// TIA Portal project "MCP_RB001002" (V15.1)

(* hardware
DEVICE "S7-1200 station_1"  S7-1200 Station
   slot 0: "Rack_0"  S7-1200 Rack  Rack  V1.0
   slot 1: "MCP"  CPU 1215C DC/DC/DC  6ES7 215-1AG40-0XB0  V4.2
DEVICE "GSD device_1"  GSD.Device.PN
   slot 0: "机架"  Rack  V1.0
   slot 0: "PNMB-address"  PNM02 V1.5  PNMB  V1.50
      slot 0: "PNM02 V1.5"  PNM02 V1.5
      slot 1: "PN-IO"  PN-IO
         slot 1: "Port 1"  Port 1
         slot 2: "Port 2"  Port 2
   slot 1: "M: 03 Read 050 Words (4xxxx)_1"  M: 03 Read 050 Words (4xxxx)
      slot 0: "M: 03 Read 050 Words (4xxxx)"  M: 03 Read 050 Words (4xxxx)
   slot 2: "M: 03 Read 050 Words (4xxxx)_2"  M: 03 Read 050 Words (4xxxx)
      slot 0: "M: 03 Read 050 Words (4xxxx)"  M: 03 Read 050 Words (4xxxx)
   slot 3: "M: 03 Read 050 Words (4xxxx)_3"  M: 03 Read 050 Words (4xxxx)
      slot 0: "M: 03 Read 050 Words (4xxxx)"  M: 03 Read 050 Words (4xxxx)
   slot 4: "M: 03 Read 050 Words (4xxxx)_4"  M: 03 Read 050 Words (4xxxx)
      slot 0: "M: 03 Read 050 Words (4xxxx)"  M: 03 Read 050 Words (4xxxx)
   slot 5: "M: 03 Read 050 Words (4xxxx)_5"  M: 03 Read 050 Words (4xxxx)
      slot 0: "M: 03 Read 050 Words (4xxxx)"  M: 03 Read 050 Words (4xxxx)
   slot 6: "M: 03 Read 002 Words (4xxxx)_1"  M: 03 Read 002 Words (4xxxx)
      slot 0: "M: 03 Read 002 Words (4xxxx)"  M: 03 Read 002 Words (4xxxx)
   slot 7: "M: 03 Read 002 Words (4xxxx)_2"  M: 03 Read 002 Words (4xxxx)
      slot 0: "M: 03 Read 002 Words (4xxxx)"  M: 03 Read 002 Words (4xxxx)
DEVICE "PC-System_1"  SIMATIC PC station
   slot 0: "SIMATIC PC station"  Rail  SIMATIC PC-Station  V1.0
      slot 125: "Stationmanager"  Station_Manager  V6.0.4
   slot 1: "IE general_1"  IE General  IE_CP  V8.2.0
   slot 2: "HMI_RT_1"  WinCC RT Advanced  6AV2 104-0xxxx-xxxx  15.1.0.0
      slot 33792: "主机接口"  Host interface
*)

// ===== PLC "MCP"  CPU 1215C DC/DC/DC =====

VAR_GLOBAL   // PLC tag table "默认变量表"
   "ID_100" AT %ID100 : Real;
   "ID_104" AT %ID104 : Real;
   "ID_108" AT %ID108 : Real;
   "ID_112" AT %ID112 : Real;
   "ID_116" AT %ID116 : Real;
   "ID_120" AT %ID120 : Real;
   "ID_124" AT %ID124 : Real;
   "ID_128" AT %ID128 : Real;
   "ID_132" AT %ID132 : Real;
   "ID_136" AT %ID136 : DInt;
   "ID_140" AT %ID140 : DInt;
   "ID_144" AT %ID144 : Real;
   "Tag_8" AT %ID148 : Real;
   "Tag_8(1)" AT %ID152 : Real;
   "Tag_9" AT %ID156 : Real;
   "ID_160" AT %IW160 : Word;
   "Tag_10" AT %ID164 : Real;
   "Tag_10(1)" AT %ID168 : Real;
   "Tag_11" AT %ID172 : Real;
   "Tag_11(1)" AT %ID176 : Real;
   "Tag_12" AT %ID180 : Real;
   "Tag_12(1)" AT %ID184 : Real;
   "Tag_13" AT %ID188 : Real;
   "Tag_13(1)" AT %ID192 : Real;
   "Tag_14" AT %ID196 : Real;
   "Tag_14(1)" AT %ID200 : Real;
   "Tag_15" AT %ID204 : Real;
   "Tag_16" AT %ID208 : Real;
   "Tag_17" AT %ID212 : Real;
   "Tag_18" AT %ID216 : Real;
   "Tag_19" AT %ID220 : Real;
   "Tag_20" AT %IW224 : Int;
   "Tag_21" AT %ID228 : Real;
   "Tag_22" AT %ID232 : Real;
   "Tag_23" AT %ID236 : Real;
   "Tag_24" AT %ID240 : Real;
   "Tag_25" AT %ID244 : Real;
   "Tag_26" AT %ID248 : Real;
   "Tag_27" AT %ID252 : Real;
   "Tag_28" AT %ID256 : Real;
   "Tag_29" AT %ID260 : Real;
   "Tag_30" AT %ID264 : Real;
   "Tag_31" AT %ID268 : Real;
   "Tag_32" AT %ID272 : Real;
   "Tag_33" AT %ID276 : Real;
   "ID_148" AT %ID148 : DWord;
   "ID_152" AT %ID152 : DWord;
   "ID_156" AT %ID156 : DWord;
   "ID_162" AT %IW162 : Word;
   "ID_164" AT %IW164 : Word;
   "ID_166" AT %IW166 : Word;
   "ID_168" AT %IW168 : Word;
   "ID_170" AT %IW170 : Word;
   "ID_172" AT %IW172 : Word;
   "ID_174" AT %IW174 : Word;
   "ID_176" AT %IW176 : Word;
   "ID_178" AT %IW178 : Word;
   "ID_180" AT %IW180 : Word;
   "ID_182" AT %IW182 : Word;
   "ID_184" AT %IW184 : Word;
   "ID_186" AT %IW186 : Word;
   "ID_188" AT %IW188 : Word;
   "ID_190" AT %IW190 : Word;
   "ID_192" AT %IW192 : Word;
   "ID_194" AT %IW194 : Word;
   "ID_196" AT %IW196 : Word;
   "ID_198" AT %IW198 : Word;
   "ID_158" AT %IW158 : Word;
   "Tag_1" AT %IW64 : Word;
   "Tag_2" AT %M100.0 : Bool;
   "Tag_3" AT %M100.1 : Bool;
   "Tag_4" AT %IW66 : Word;
   "Tag_5" AT %ID600 : DInt;
   "Tag_6" AT %ID700 : DInt;
   "Tag_7" AT %MD104 : DInt;
   "Tag_34" AT %MD108 : DInt;
   "System_Byte" AT %MB1 : Byte;
   "FirstScan" AT %M1.0 : Bool;
   "DiagStatusUpdate" AT %M1.1 : Bool;
   "AlwaysTRUE" AT %M1.2 : Bool;
   "AlwaysFALSE" AT %M1.3 : Bool;
   "Clock_Byte" AT %MB0 : Byte;
   "Clock_10Hz" AT %M0.0 : Bool;
   "Clock_5Hz" AT %M0.1 : Bool;
   "Clock_2.5Hz" AT %M0.2 : Bool;
   "Clock_2Hz" AT %M0.3 : Bool;
   "Clock_1.25Hz" AT %M0.4 : Bool;
   "Clock_1Hz" AT %M0.5 : Bool;
   "Clock_0.625Hz" AT %M0.6 : Bool;
   "Clock_0.5Hz" AT %M0.7 : Bool;
   "Tag_35" AT %M100.2 : Bool;
END_VAR

VAR_GLOBAL   // PLC tag table "精炼机采集"
   "N11" AT %I100.0 : "精炼机";
   "N12" AT %I200.0 : "精炼机";
   "N13" AT %I300.0 : "精炼机";
   "N14" AT %I400.0 : "精炼机";
   "N15" AT %I500.0 : "精炼机";
END_VAR

TYPE "精炼机"
   STRUCT
      左前辊温度 : Real;
      右前辊温度 : Real;
      左后辊温度 : Real;
      右后辊温度 : Real;
      左间隙 : Real;
      右间隙 : Real;
      滚筒电机电流 : Real;
      滚筒电机频率 : Real;
      滚筒电机功率 : Real;
      滚筒电机电度 : DInt;
      滚筒电机计时 : DInt;
      环境温度 : Real;
      环境湿度 : Real;
      胶温 : Real;
      开关量汇总 : DInt;
      当前任务编号 : Array[0..9] of WChar;
      当前人员编号 : Array[0..9] of WChar;
   END_STRUCT;
END_TYPE

TYPE "精炼机上传"
   STRUCT
      左前辊温度 : Real;
      右前辊温度 : Real;
      左后辊温度 : Real;
      右后辊温度 : Real;
      左间隙 : Real;
      右间隙 : Real;
      滚筒电机电流 : Real;
      滚筒电机频率 : Real;
      滚筒电机功率 : Real;
      滚筒电机电度 : DInt;
      滚筒电机计时 : DInt;
      环境温度 : Real;
      环境湿度 : Real;
      胶温 : Real;
      开关量汇总 : DInt;
      当前任务编号 : Array[0..9] of WChar;
      当前人员编号 : Array[0..9] of WChar;
   END_STRUCT;
END_TYPE

TYPE "uMySQL_CDD"
   STRUCT
      Connect_OK : Bool;
      Connect_ID : Conn_Ouc;
      Connect_Sequence : DInt;
      Server_Protocol_Version : Int;
      Server_Server_Version : String;
      Server_Character_Set : Byte;
      CLIENT_PLUGIN_AUTH : String;
      Recv_Done : Bool;
      Recv_Len : Int;
      Recv_Buffer : Array[0..2048] of Byte;
      Send_Done : Bool;
      Send_Len : Int;
      Send_Buffer : Array[0..2048] of Byte;
   END_STRUCT;
END_TYPE

TYPE "精炼机数据库"
   STRUCT
      左前辊温度 : Real;
      右前辊温度 : Real;
      左后辊温度 : Real;
      右后辊温度 : Real;
      左间隙 : Real;
      右间隙 : Real;
      滚筒电机电流 : Real;
      滚筒电机频率 : Real;
      滚筒电机功率 : Real;
      滚筒电机电度 : DInt;
      滚筒电机计时 : DInt;
      环境温度 : Real;
      环境湿度 : Real;
      胶温 : Real;
      开关量汇总 : DInt;
      当前任务编号 : WString;
      当前人员编号 : WString;
   END_STRUCT;
END_TYPE

DATA_BLOCK "精炼机数据转存"   // DB100
{ S7_Optimized_Access := 'FALSE' }
VERSION : 0.1
   VAR
      Temp : Array[0..99] of Byte;
      N11精炼机 : "精炼机上传";
      N12精炼机 : "精炼机上传";
      N13精炼机 : "精炼机上传";
      N14精炼机 : "精炼机上传";
      N15精炼机 : "精炼机上传";
      N21卷片机累计重量 : DInt;
      N22卷片机累计重量 : DInt;
   END_VAR
BEGIN
END_DATA_BLOCK

DATA_BLOCK "通用数据采集"   // DB200
{ S7_Optimized_Access := 'TRUE' }
VERSION : 0.1
   VAR
      环境温度 : Real;
      环境湿度 : Real;
   END_VAR
BEGIN
END_DATA_BLOCK

DATA_BLOCK "温控相机解码_N15"   // DB405
{ S7_Optimized_Access := 'TRUE' }
VERSION : 0.1
// stored: InstanceOfName 温控相机解码
"温控相机解码"
BEGIN
END_DATA_BLOCK

// folder: System blocks/Program resources

DATA_BLOCK "IEC_Timer_0_DB"   // DB1
{ S7_Optimized_Access := 'TRUE' }
AUTHOR : Simatic
FAMILY : IEC
NAME : IEC_TMR
VERSION : 1.0
// stored: InstanceOfName IEC_TIMER
"IEC_TIMER"
BEGIN
END_DATA_BLOCK

// folder: 存数据库

DATA_BLOCK "Wchartest"   // DB2
{ S7_Optimized_Access := 'TRUE' }
VERSION : 0.1
   VAR
      TemWchar : WChar;
      TemWstring : WString;
      WstringLen : UInt;
      ArrayWCHAR : Array[0..1023] of WChar;
      ArrayChar : Array[0..1023] of Char;
      arraayWord : Array[0..1023] of Word;
   END_VAR
BEGIN
END_DATA_BLOCK

DATA_BLOCK "数据库字符串"   // DB900
{ S7_Optimized_Access := 'TRUE' }
VERSION : 0.1
   VAR
      wstring : WString[2048];
   END_VAR
   VAR RETAIN
      Connect_CMD : Bool;
   END_VAR
   VAR
      Connect_CND : Bool;
      Connect_Error : Bool;
      Use_CMD : Bool;
      Use_Done : Bool;
      Use_Error : Bool;
      Query_CMD : Bool;
      Query_Done : Bool;
      Query_Error : Bool;
      CommandLine : WString[2048];
   END_VAR
   VAR RETAIN
      SerialNum : Int := 1;
   END_VAR
   VAR
      Addr : Int := 11;
      UploadData : "精炼机数据库";
      Upload : Array[11..15] of "精炼机数据库";
   END_VAR
BEGIN
END_DATA_BLOCK

DATA_BLOCK "uMySQL_Connect_DB"   // DB901
{ S7_Optimized_Access := 'TRUE' }
VERSION : 0.1
// stored: InstanceOfName uMySQL_Connect
"uMySQL_Connect"
BEGIN
   IP.RemoteAddress.ADDR[3] := 16#A0;
   IP.RemoteAddress.ADDR[4] := 16#A3;
   Net_ID := 16#0070;
   UserName := 'plc';
   DB_Name := 'rb001011';
   IP.InterfaceId := 64;
   IP.ID := 16#0070;
   IP.ConnectionType := 16#0B;
   IP.ActiveEstablished := TRUE;
   TempBool[1] := TRUE;
   SND_Buffer[0] := 16#01;
   SND_Buffer[4] := 16#01;
   NetConnect.STATUS := 16#7000;
   NetRcv.ADHOC := TRUE;
   NetRcv.STATUS := 16#7000;
   "Step" := 6;
   ServerCapability_flag := 16#0000_0000;
   Client_CapabilityFlag := 16#0000_8609;
   Client_MaxLen := 16#0000_0000;
   NetDISCON.ID := 16#0070;
   NetDISCON.STATUS := 16#7000;
   NetSend.ID := 16#0070;
   NetSend.STATUS := 16#7000;
   NetDiag.REQ := TRUE;
   NetDiag.ID := 16#0070;
   NetDiag.BUSY := TRUE;
   NetDiag.STATUS := 16#7001;
   Timer_ON.ST := T#10D_22H_43M_20S_90MS;
   Timer_ON.PT := T#500MS;
   Timer_ON.RU := TRUE;
   Timer_ON.IN := TRUE;
   Timer_OFF.ST := T#10D_22H_43M_19S_563MS;
   Timer_OFF.PT := T#500MS;
   NetSendEnd.REQ := TRUE;
   NetSendEnd.ID := 16#0070;
   NetSendEnd.LEN := 5;
   NetSendEnd.STATUS := 16#7000;
   NetSendEnd_EN := TRUE;
   SendWChar[0] := WCHAR#' ';
   SendWChar[1] := WCHAR#' ';
   SendWChar[2] := WCHAR#' ';
   SendWChar[3] := WCHAR#' ';
   SendWChar[4] := WCHAR#' ';
   SendWChar[5] := WCHAR#' ';
   SendWChar[6] := WCHAR#' ';
   SendWChar[7] := WCHAR#' ';
   SendWChar[8] := WCHAR#' ';
   SendWChar[9] := WCHAR#' ';
   SendWChar[10] := WCHAR#' ';
   SendWChar[11] := WCHAR#' ';
   SendWChar[12] := WCHAR#' ';
   SendWChar[13] := WCHAR#' ';
   SendWChar[14] := WCHAR#' ';
   SendWChar[15] := WCHAR#' ';
   SendWChar[16] := WCHAR#' ';
   SendWChar[17] := WCHAR#' ';
   SendWChar[18] := WCHAR#' ';
   SendWChar[19] := WCHAR#' ';
   SendWChar[20] := WCHAR#' ';
   SendWChar[21] := WCHAR#' ';
   SendWChar[22] := WCHAR#' ';
   SendWChar[23] := WCHAR#' ';
   SendWChar[24] := WCHAR#' ';
   SendWChar[25] := WCHAR#' ';
   SendWChar[26] := WCHAR#' ';
   SendWChar[27] := WCHAR#' ';
   SendWChar[28] := WCHAR#' ';
   SendWChar[29] := WCHAR#' ';
   SendWChar[30] := WCHAR#' ';
   SendWChar[31] := WCHAR#' ';
   SendWChar[32] := WCHAR#' ';
   SendWChar[33] := WCHAR#' ';
   SendWChar[34] := WCHAR#' ';
   SendWChar[35] := WCHAR#' ';
   SendWChar[36] := WCHAR#' ';
   SendWChar[37] := WCHAR#' ';
   SendWChar[38] := WCHAR#' ';
   SendWChar[39] := WCHAR#' ';
   SendWChar[40] := WCHAR#' ';
   SendWChar[41] := WCHAR#' ';
   SendWChar[42] := WCHAR#' ';
   SendWChar[43] := WCHAR#' ';
   SendWChar[44] := WCHAR#' ';
   SendWChar[45] := WCHAR#' ';
   SendWChar[46] := WCHAR#' ';
   SendWChar[47] := WCHAR#' ';
   SendWChar[48] := WCHAR#' ';
   SendWChar[49] := WCHAR#' ';
   SendWChar[50] := WCHAR#' ';
   SendWChar[51] := WCHAR#' ';
   SendWChar[52] := WCHAR#' ';
   SendWChar[53] := WCHAR#' ';
   SendWChar[54] := WCHAR#' ';
   SendWChar[55] := WCHAR#' ';
   SendWChar[56] := WCHAR#' ';
   SendWChar[57] := WCHAR#' ';
   SendWChar[58] := WCHAR#' ';
   SendWChar[59] := WCHAR#' ';
   SendWChar[60] := WCHAR#' ';
   SendWChar[61] := WCHAR#' ';
   SendWChar[62] := WCHAR#' ';
   SendWChar[63] := WCHAR#' ';
   SendWChar[64] := WCHAR#' ';
   SendWChar[65] := WCHAR#' ';
   SendWChar[66] := WCHAR#' ';
   SendWChar[67] := WCHAR#' ';
   SendWChar[68] := WCHAR#' ';
   SendWChar[69] := WCHAR#' ';
   SendWChar[70] := WCHAR#' ';
   SendWChar[71] := WCHAR#' ';
   SendWChar[72] := WCHAR#' ';
   SendWChar[73] := WCHAR#' ';
   SendWChar[74] := WCHAR#' ';
   SendWChar[75] := WCHAR#' ';
   SendWChar[76] := WCHAR#' ';
   SendWChar[77] := WCHAR#' ';
   SendWChar[78] := WCHAR#' ';
   SendWChar[79] := WCHAR#' ';
   SendWChar[80] := WCHAR#' ';
   SendWChar[81] := WCHAR#' ';
   SendWChar[82] := WCHAR#' ';
   SendWChar[83] := WCHAR#' ';
   SendWChar[84] := WCHAR#' ';
   SendWChar[85] := WCHAR#' ';
   SendWChar[86] := WCHAR#' ';
   SendWChar[87] := WCHAR#' ';
   SendWChar[88] := WCHAR#' ';
   SendWChar[89] := WCHAR#' ';
   SendWChar[90] := WCHAR#' ';
   SendWChar[91] := WCHAR#' ';
   SendWChar[92] := WCHAR#' ';
   SendWChar[93] := WCHAR#' ';
   SendWChar[94] := WCHAR#' ';
   SendWChar[95] := WCHAR#' ';
   SendWChar[96] := WCHAR#' ';
   SendWChar[97] := WCHAR#' ';
   SendWChar[98] := WCHAR#' ';
   SendWChar[99] := WCHAR#' ';
   SendWChar[100] := WCHAR#' ';
   SendWChar[101] := WCHAR#' ';
   SendWChar[102] := WCHAR#' ';
   SendWChar[103] := WCHAR#' ';
   SendWChar[104] := WCHAR#' ';
   SendWChar[105] := WCHAR#' ';
   SendWChar[106] := WCHAR#' ';
   SendWChar[107] := WCHAR#' ';
   SendWChar[108] := WCHAR#' ';
   SendWChar[109] := WCHAR#' ';
   SendWChar[110] := WCHAR#' ';
   SendWChar[111] := WCHAR#' ';
   SendWChar[112] := WCHAR#' ';
   SendWChar[113] := WCHAR#' ';
   SendWChar[114] := WCHAR#' ';
   SendWChar[115] := WCHAR#' ';
   SendWChar[116] := WCHAR#' ';
   SendWChar[117] := WCHAR#' ';
   SendWChar[118] := WCHAR#' ';
   SendWChar[119] := WCHAR#' ';
   SendWChar[120] := WCHAR#' ';
   SendWChar[121] := WCHAR#' ';
   SendWChar[122] := WCHAR#' ';
   SendWChar[123] := WCHAR#' ';
   SendWChar[124] := WCHAR#' ';
   SendWChar[125] := WCHAR#' ';
   SendWChar[126] := WCHAR#' ';
   SendWChar[127] := WCHAR#' ';
   SendWChar[128] := WCHAR#' ';
   SendWChar[129] := WCHAR#' ';
   SendWChar[130] := WCHAR#' ';
   SendWChar[131] := WCHAR#' ';
   SendWChar[132] := WCHAR#' ';
   SendWChar[133] := WCHAR#' ';
   SendWChar[134] := WCHAR#' ';
   SendWChar[135] := WCHAR#' ';
   SendWChar[136] := WCHAR#' ';
   SendWChar[137] := WCHAR#' ';
   SendWChar[138] := WCHAR#' ';
   SendWChar[139] := WCHAR#' ';
   SendWChar[140] := WCHAR#' ';
   SendWChar[141] := WCHAR#' ';
   SendWChar[142] := WCHAR#' ';
   SendWChar[143] := WCHAR#' ';
   SendWChar[144] := WCHAR#' ';
   SendWChar[145] := WCHAR#' ';
   SendWChar[146] := WCHAR#' ';
   SendWChar[147] := WCHAR#' ';
   SendWChar[148] := WCHAR#' ';
   SendWChar[149] := WCHAR#' ';
   SendWChar[150] := WCHAR#' ';
   SendWChar[151] := WCHAR#' ';
   SendWChar[152] := WCHAR#' ';
   SendWChar[153] := WCHAR#' ';
   SendWChar[154] := WCHAR#' ';
   SendWChar[155] := WCHAR#' ';
   SendWChar[156] := WCHAR#' ';
   SendWChar[157] := WCHAR#' ';
   SendWChar[158] := WCHAR#' ';
   SendWChar[159] := WCHAR#' ';
   SendWChar[160] := WCHAR#' ';
   SendWChar[161] := WCHAR#' ';
   SendWChar[162] := WCHAR#' ';
   SendWChar[163] := WCHAR#' ';
   SendWChar[164] := WCHAR#' ';
   SendWChar[165] := WCHAR#' ';
   SendWChar[166] := WCHAR#' ';
   SendWChar[167] := WCHAR#' ';
   SendWChar[168] := WCHAR#' ';
   SendWChar[169] := WCHAR#' ';
   SendWChar[170] := WCHAR#' ';
   SendWChar[171] := WCHAR#' ';
   SendWChar[172] := WCHAR#' ';
   SendWChar[173] := WCHAR#' ';
   SendWChar[174] := WCHAR#' ';
   SendWChar[175] := WCHAR#' ';
   SendWChar[176] := WCHAR#' ';
   SendWChar[177] := WCHAR#' ';
   SendWChar[178] := WCHAR#' ';
   SendWChar[179] := WCHAR#' ';
   SendWChar[180] := WCHAR#' ';
   SendWChar[181] := WCHAR#' ';
   SendWChar[182] := WCHAR#' ';
   SendWChar[183] := WCHAR#' ';
   SendWChar[184] := WCHAR#' ';
   SendWChar[185] := WCHAR#' ';
   SendWChar[186] := WCHAR#' ';
   SendWChar[187] := WCHAR#' ';
   SendWChar[188] := WCHAR#' ';
   SendWChar[189] := WCHAR#' ';
   SendWChar[190] := WCHAR#' ';
   SendWChar[191] := WCHAR#' ';
   SendWChar[192] := WCHAR#' ';
   SendWChar[193] := WCHAR#' ';
   SendWChar[194] := WCHAR#' ';
   SendWChar[195] := WCHAR#' ';
   SendWChar[196] := WCHAR#' ';
   SendWChar[197] := WCHAR#' ';
   SendWChar[198] := WCHAR#' ';
   SendWChar[199] := WCHAR#' ';
   SendWChar[200] := WCHAR#' ';
   SendWChar[201] := WCHAR#' ';
   SendWChar[202] := WCHAR#' ';
   SendWChar[203] := WCHAR#' ';
   SendWChar[204] := WCHAR#' ';
   SendWChar[205] := WCHAR#' ';
   SendWChar[206] := WCHAR#' ';
   SendWChar[207] := WCHAR#' ';
   SendWChar[208] := WCHAR#' ';
   SendWChar[209] := WCHAR#' ';
   SendWChar[210] := WCHAR#' ';
   SendWChar[211] := WCHAR#' ';
   SendWChar[212] := WCHAR#' ';
   SendWChar[213] := WCHAR#' ';
   SendWChar[214] := WCHAR#' ';
   SendWChar[215] := WCHAR#' ';
   SendWChar[216] := WCHAR#' ';
   SendWChar[217] := WCHAR#' ';
   SendWChar[218] := WCHAR#' ';
   SendWChar[219] := WCHAR#' ';
   SendWChar[220] := WCHAR#' ';
   SendWChar[221] := WCHAR#' ';
   SendWChar[222] := WCHAR#' ';
   SendWChar[223] := WCHAR#' ';
   SendWChar[224] := WCHAR#' ';
   SendWChar[225] := WCHAR#' ';
   SendWChar[226] := WCHAR#' ';
   SendWChar[227] := WCHAR#' ';
   SendWChar[228] := WCHAR#' ';
   SendWChar[229] := WCHAR#' ';
   SendWChar[230] := WCHAR#' ';
   SendWChar[231] := WCHAR#' ';
   SendWChar[232] := WCHAR#' ';
   SendWChar[233] := WCHAR#' ';
   SendWChar[234] := WCHAR#' ';
   SendWChar[235] := WCHAR#' ';
   SendWChar[236] := WCHAR#' ';
   SendWChar[237] := WCHAR#' ';
   SendWChar[238] := WCHAR#' ';
   SendWChar[239] := WCHAR#' ';
   SendWChar[240] := WCHAR#' ';
   SendWChar[241] := WCHAR#' ';
   SendWChar[242] := WCHAR#' ';
   SendWChar[243] := WCHAR#' ';
   SendWChar[244] := WCHAR#' ';
   SendWChar[245] := WCHAR#' ';
   SendWChar[246] := WCHAR#' ';
   SendWChar[247] := WCHAR#' ';
   SendWChar[248] := WCHAR#' ';
   SendWChar[249] := WCHAR#' ';
   SendWChar[250] := WCHAR#' ';
   SendWChar[251] := WCHAR#' ';
   SendWChar[252] := WCHAR#' ';
   SendWChar[253] := WCHAR#' ';
   SendWChar[254] := WCHAR#' ';
   SendWChar[255] := WCHAR#' ';
   SendWChar[256] := WCHAR#' ';
   SendWChar[257] := WCHAR#' ';
   SendWChar[258] := WCHAR#' ';
   SendWChar[259] := WCHAR#' ';
   SendWChar[260] := WCHAR#' ';
   SendWChar[261] := WCHAR#' ';
   SendWChar[262] := WCHAR#' ';
   SendWChar[263] := WCHAR#' ';
   SendWChar[264] := WCHAR#' ';
   SendWChar[265] := WCHAR#' ';
   SendWChar[266] := WCHAR#' ';
   SendWChar[267] := WCHAR#' ';
   SendWChar[268] := WCHAR#' ';
   SendWChar[269] := WCHAR#' ';
   SendWChar[270] := WCHAR#' ';
   SendWChar[271] := WCHAR#' ';
   SendWChar[272] := WCHAR#' ';
   SendWChar[273] := WCHAR#' ';
   SendWChar[274] := WCHAR#' ';
   SendWChar[275] := WCHAR#' ';
   SendWChar[276] := WCHAR#' ';
   SendWChar[277] := WCHAR#' ';
   SendWChar[278] := WCHAR#' ';
   SendWChar[279] := WCHAR#' ';
   SendWChar[280] := WCHAR#' ';
   SendWChar[281] := WCHAR#' ';
   SendWChar[282] := WCHAR#' ';
   SendWChar[283] := WCHAR#' ';
   SendWChar[284] := WCHAR#' ';
   SendWChar[285] := WCHAR#' ';
   SendWChar[286] := WCHAR#' ';
   SendWChar[287] := WCHAR#' ';
   SendWChar[288] := WCHAR#' ';
   SendWChar[289] := WCHAR#' ';
   SendWChar[290] := WCHAR#' ';
   SendWChar[291] := WCHAR#' ';
   SendWChar[292] := WCHAR#' ';
   SendWChar[293] := WCHAR#' ';
   SendWChar[294] := WCHAR#' ';
   SendWChar[295] := WCHAR#' ';
   SendWChar[296] := WCHAR#' ';
   SendWChar[297] := WCHAR#' ';
   SendWChar[298] := WCHAR#' ';
   SendWChar[299] := WCHAR#' ';
   SendWChar[300] := WCHAR#' ';
   SendWChar[301] := WCHAR#' ';
   SendWChar[302] := WCHAR#' ';
   SendWChar[303] := WCHAR#' ';
   SendWChar[304] := WCHAR#' ';
   SendWChar[305] := WCHAR#' ';
   SendWChar[306] := WCHAR#' ';
   SendWChar[307] := WCHAR#' ';
   SendWChar[308] := WCHAR#' ';
   SendWChar[309] := WCHAR#' ';
   SendWChar[310] := WCHAR#' ';
   SendWChar[311] := WCHAR#' ';
   SendWChar[312] := WCHAR#' ';
   SendWChar[313] := WCHAR#' ';
   SendWChar[314] := WCHAR#' ';
   SendWChar[315] := WCHAR#' ';
   SendWChar[316] := WCHAR#' ';
   SendWChar[317] := WCHAR#' ';
   SendWChar[318] := WCHAR#' ';
   SendWChar[319] := WCHAR#' ';
   SendWChar[320] := WCHAR#' ';
   SendWChar[321] := WCHAR#' ';
   SendWChar[322] := WCHAR#' ';
   SendWChar[323] := WCHAR#' ';
   SendWChar[324] := WCHAR#' ';
   SendWChar[325] := WCHAR#' ';
   SendWChar[326] := WCHAR#' ';
   SendWChar[327] := WCHAR#' ';
   SendWChar[328] := WCHAR#' ';
   SendWChar[329] := WCHAR#' ';
   SendWChar[330] := WCHAR#' ';
   SendWChar[331] := WCHAR#' ';
   SendWChar[332] := WCHAR#' ';
   SendWChar[333] := WCHAR#' ';
   SendWChar[334] := WCHAR#' ';
   SendWChar[335] := WCHAR#' ';
   SendWChar[336] := WCHAR#' ';
   SendWChar[337] := WCHAR#' ';
   SendWChar[338] := WCHAR#' ';
   SendWChar[339] := WCHAR#' ';
   SendWChar[340] := WCHAR#' ';
   SendWChar[341] := WCHAR#' ';
   SendWChar[342] := WCHAR#' ';
   SendWChar[343] := WCHAR#' ';
   SendWChar[344] := WCHAR#' ';
   SendWChar[345] := WCHAR#' ';
   SendWChar[346] := WCHAR#' ';
   SendWChar[347] := WCHAR#' ';
   SendWChar[348] := WCHAR#' ';
   SendWChar[349] := WCHAR#' ';
   SendWChar[350] := WCHAR#' ';
   SendWChar[351] := WCHAR#' ';
   SendWChar[352] := WCHAR#' ';
   SendWChar[353] := WCHAR#' ';
   SendWChar[354] := WCHAR#' ';
   SendWChar[355] := WCHAR#' ';
   SendWChar[356] := WCHAR#' ';
   SendWChar[357] := WCHAR#' ';
   SendWChar[358] := WCHAR#' ';
   SendWChar[359] := WCHAR#' ';
   SendWChar[360] := WCHAR#' ';
   SendWChar[361] := WCHAR#' ';
   SendWChar[362] := WCHAR#' ';
   SendWChar[363] := WCHAR#' ';
   SendWChar[364] := WCHAR#' ';
   SendWChar[365] := WCHAR#' ';
   SendWChar[366] := WCHAR#' ';
   SendWChar[367] := WCHAR#' ';
   SendWChar[368] := WCHAR#' ';
   SendWChar[369] := WCHAR#' ';
   SendWChar[370] := WCHAR#' ';
   SendWChar[371] := WCHAR#' ';
   SendWChar[372] := WCHAR#' ';
   SendWChar[373] := WCHAR#' ';
   SendWChar[374] := WCHAR#' ';
   SendWChar[375] := WCHAR#' ';
   SendWChar[376] := WCHAR#' ';
   SendWChar[377] := WCHAR#' ';
   SendWChar[378] := WCHAR#' ';
   SendWChar[379] := WCHAR#' ';
   SendWChar[380] := WCHAR#' ';
   SendWChar[381] := WCHAR#' ';
   SendWChar[382] := WCHAR#' ';
   SendWChar[383] := WCHAR#' ';
   SendWChar[384] := WCHAR#' ';
   SendWChar[385] := WCHAR#' ';
   SendWChar[386] := WCHAR#' ';
   SendWChar[387] := WCHAR#' ';
   SendWChar[388] := WCHAR#' ';
   SendWChar[389] := WCHAR#' ';
   SendWChar[390] := WCHAR#' ';
   SendWChar[391] := WCHAR#' ';
   SendWChar[392] := WCHAR#' ';
   SendWChar[393] := WCHAR#' ';
   SendWChar[394] := WCHAR#' ';
   SendWChar[395] := WCHAR#' ';
   SendWChar[396] := WCHAR#' ';
   SendWChar[397] := WCHAR#' ';
   SendWChar[398] := WCHAR#' ';
   SendWChar[399] := WCHAR#' ';
   SendWChar[400] := WCHAR#' ';
   SendWChar[401] := WCHAR#' ';
   SendWChar[402] := WCHAR#' ';
   SendWChar[403] := WCHAR#' ';
   SendWChar[404] := WCHAR#' ';
   SendWChar[405] := WCHAR#' ';
   SendWChar[406] := WCHAR#' ';
   SendWChar[407] := WCHAR#' ';
   SendWChar[408] := WCHAR#' ';
   SendWChar[409] := WCHAR#' ';
   SendWChar[410] := WCHAR#' ';
   SendWChar[411] := WCHAR#' ';
   SendWChar[412] := WCHAR#' ';
   SendWChar[413] := WCHAR#' ';
   SendWChar[414] := WCHAR#' ';
   SendWChar[415] := WCHAR#' ';
   SendWChar[416] := WCHAR#' ';
   SendWChar[417] := WCHAR#' ';
   SendWChar[418] := WCHAR#' ';
   SendWChar[419] := WCHAR#' ';
   SendWChar[420] := WCHAR#' ';
   SendWChar[421] := WCHAR#' ';
   SendWChar[422] := WCHAR#' ';
   SendWChar[423] := WCHAR#' ';
   SendWChar[424] := WCHAR#' ';
   SendWChar[425] := WCHAR#' ';
   SendWChar[426] := WCHAR#' ';
   SendWChar[427] := WCHAR#' ';
   SendWChar[428] := WCHAR#' ';
   SendWChar[429] := WCHAR#' ';
   SendWChar[430] := WCHAR#' ';
   SendWChar[431] := WCHAR#' ';
   SendWChar[432] := WCHAR#' ';
   SendWChar[433] := WCHAR#' ';
   SendWChar[434] := WCHAR#' ';
   SendWChar[435] := WCHAR#' ';
   SendWChar[436] := WCHAR#' ';
   SendWChar[437] := WCHAR#' ';
   SendWChar[438] := WCHAR#' ';
   SendWChar[439] := WCHAR#' ';
   SendWChar[440] := WCHAR#' ';
   SendWChar[441] := WCHAR#' ';
   SendWChar[442] := WCHAR#' ';
   SendWChar[443] := WCHAR#' ';
   SendWChar[444] := WCHAR#' ';
   SendWChar[445] := WCHAR#' ';
   SendWChar[446] := WCHAR#' ';
   SendWChar[447] := WCHAR#' ';
   SendWChar[448] := WCHAR#' ';
   SendWChar[449] := WCHAR#' ';
   SendWChar[450] := WCHAR#' ';
   SendWChar[451] := WCHAR#' ';
   SendWChar[452] := WCHAR#' ';
   SendWChar[453] := WCHAR#' ';
   SendWChar[454] := WCHAR#' ';
   SendWChar[455] := WCHAR#' ';
   SendWChar[456] := WCHAR#' ';
   SendWChar[457] := WCHAR#' ';
   SendWChar[458] := WCHAR#' ';
   SendWChar[459] := WCHAR#' ';
   SendWChar[460] := WCHAR#' ';
   SendWChar[461] := WCHAR#' ';
   SendWChar[462] := WCHAR#' ';
   SendWChar[463] := WCHAR#' ';
   SendWChar[464] := WCHAR#' ';
   SendWChar[465] := WCHAR#' ';
   SendWChar[466] := WCHAR#' ';
   SendWChar[467] := WCHAR#' ';
   SendWChar[468] := WCHAR#' ';
   SendWChar[469] := WCHAR#' ';
   SendWChar[470] := WCHAR#' ';
   SendWChar[471] := WCHAR#' ';
   SendWChar[472] := WCHAR#' ';
   SendWChar[473] := WCHAR#' ';
   SendWChar[474] := WCHAR#' ';
   SendWChar[475] := WCHAR#' ';
   SendWChar[476] := WCHAR#' ';
   SendWChar[477] := WCHAR#' ';
   SendWChar[478] := WCHAR#' ';
   SendWChar[479] := WCHAR#' ';
   SendWChar[480] := WCHAR#' ';
   SendWChar[481] := WCHAR#' ';
   SendWChar[482] := WCHAR#' ';
   SendWChar[483] := WCHAR#' ';
   SendWChar[484] := WCHAR#' ';
   SendWChar[485] := WCHAR#' ';
   SendWChar[486] := WCHAR#' ';
   SendWChar[487] := WCHAR#' ';
   SendWChar[488] := WCHAR#' ';
   SendWChar[489] := WCHAR#' ';
   SendWChar[490] := WCHAR#' ';
   SendWChar[491] := WCHAR#' ';
   SendWChar[492] := WCHAR#' ';
   SendWChar[493] := WCHAR#' ';
   SendWChar[494] := WCHAR#' ';
   SendWChar[495] := WCHAR#' ';
   SendWChar[496] := WCHAR#' ';
   SendWChar[497] := WCHAR#' ';
   SendWChar[498] := WCHAR#' ';
   SendWChar[499] := WCHAR#' ';
   SendWChar[500] := WCHAR#' ';
   SendWChar[501] := WCHAR#' ';
   SendWChar[502] := WCHAR#' ';
   SendWChar[503] := WCHAR#' ';
   SendWChar[504] := WCHAR#' ';
   SendWChar[505] := WCHAR#' ';
   SendWChar[506] := WCHAR#' ';
   SendWChar[507] := WCHAR#' ';
   SendWChar[508] := WCHAR#' ';
   SendWChar[509] := WCHAR#' ';
   SendWChar[510] := WCHAR#' ';
   SendWChar[511] := WCHAR#' ';
   SendWChar[512] := WCHAR#' ';
   SendWChar[513] := WCHAR#' ';
   SendWChar[514] := WCHAR#' ';
   SendWChar[515] := WCHAR#' ';
   SendWChar[516] := WCHAR#' ';
   SendWChar[517] := WCHAR#' ';
   SendWChar[518] := WCHAR#' ';
   SendWChar[519] := WCHAR#' ';
   SendWChar[520] := WCHAR#' ';
   SendWChar[521] := WCHAR#' ';
   SendWChar[522] := WCHAR#' ';
   SendWChar[523] := WCHAR#' ';
   SendWChar[524] := WCHAR#' ';
   SendWChar[525] := WCHAR#' ';
   SendWChar[526] := WCHAR#' ';
   SendWChar[527] := WCHAR#' ';
   SendWChar[528] := WCHAR#' ';
   SendWChar[529] := WCHAR#' ';
   SendWChar[530] := WCHAR#' ';
   SendWChar[531] := WCHAR#' ';
   SendWChar[532] := WCHAR#' ';
   SendWChar[533] := WCHAR#' ';
   SendWChar[534] := WCHAR#' ';
   SendWChar[535] := WCHAR#' ';
   SendWChar[536] := WCHAR#' ';
   SendWChar[537] := WCHAR#' ';
   SendWChar[538] := WCHAR#' ';
   SendWChar[539] := WCHAR#' ';
   SendWChar[540] := WCHAR#' ';
   SendWChar[541] := WCHAR#' ';
   SendWChar[542] := WCHAR#' ';
   SendWChar[543] := WCHAR#' ';
   SendWChar[544] := WCHAR#' ';
   SendWChar[545] := WCHAR#' ';
   SendWChar[546] := WCHAR#' ';
   SendWChar[547] := WCHAR#' ';
   SendWChar[548] := WCHAR#' ';
   SendWChar[549] := WCHAR#' ';
   SendWChar[550] := WCHAR#' ';
   SendWChar[551] := WCHAR#' ';
   SendWChar[552] := WCHAR#' ';
   SendWChar[553] := WCHAR#' ';
   SendWChar[554] := WCHAR#' ';
   SendWChar[555] := WCHAR#' ';
   SendWChar[556] := WCHAR#' ';
   SendWChar[557] := WCHAR#' ';
   SendWChar[558] := WCHAR#' ';
   SendWChar[559] := WCHAR#' ';
   SendWChar[560] := WCHAR#' ';
   SendWChar[561] := WCHAR#' ';
   SendWChar[562] := WCHAR#' ';
   SendWChar[563] := WCHAR#' ';
   SendWChar[564] := WCHAR#' ';
   SendWChar[565] := WCHAR#' ';
   SendWChar[566] := WCHAR#' ';
   SendWChar[567] := WCHAR#' ';
   SendWChar[568] := WCHAR#' ';
   SendWChar[569] := WCHAR#' ';
   SendWChar[570] := WCHAR#' ';
   SendWChar[571] := WCHAR#' ';
   SendWChar[572] := WCHAR#' ';
   SendWChar[573] := WCHAR#' ';
   SendWChar[574] := WCHAR#' ';
   SendWChar[575] := WCHAR#' ';
   SendWChar[576] := WCHAR#' ';
   SendWChar[577] := WCHAR#' ';
   SendWChar[578] := WCHAR#' ';
   SendWChar[579] := WCHAR#' ';
   SendWChar[580] := WCHAR#' ';
   SendWChar[581] := WCHAR#' ';
   SendWChar[582] := WCHAR#' ';
   SendWChar[583] := WCHAR#' ';
   SendWChar[584] := WCHAR#' ';
   SendWChar[585] := WCHAR#' ';
   SendWChar[586] := WCHAR#' ';
   SendWChar[587] := WCHAR#' ';
   SendWChar[588] := WCHAR#' ';
   SendWChar[589] := WCHAR#' ';
   SendWChar[590] := WCHAR#' ';
   SendWChar[591] := WCHAR#' ';
   SendWChar[592] := WCHAR#' ';
   SendWChar[593] := WCHAR#' ';
   SendWChar[594] := WCHAR#' ';
   SendWChar[595] := WCHAR#' ';
   SendWChar[596] := WCHAR#' ';
   SendWChar[597] := WCHAR#' ';
   SendWChar[598] := WCHAR#' ';
   SendWChar[599] := WCHAR#' ';
   SendWChar[600] := WCHAR#' ';
   SendWChar[601] := WCHAR#' ';
   SendWChar[602] := WCHAR#' ';
   SendWChar[603] := WCHAR#' ';
   SendWChar[604] := WCHAR#' ';
   SendWChar[605] := WCHAR#' ';
   SendWChar[606] := WCHAR#' ';
   SendWChar[607] := WCHAR#' ';
   SendWChar[608] := WCHAR#' ';
   SendWChar[609] := WCHAR#' ';
   SendWChar[610] := WCHAR#' ';
   SendWChar[611] := WCHAR#' ';
   SendWChar[612] := WCHAR#' ';
   SendWChar[613] := WCHAR#' ';
   SendWChar[614] := WCHAR#' ';
   SendWChar[615] := WCHAR#' ';
   SendWChar[616] := WCHAR#' ';
   SendWChar[617] := WCHAR#' ';
   SendWChar[618] := WCHAR#' ';
   SendWChar[619] := WCHAR#' ';
   SendWChar[620] := WCHAR#' ';
   SendWChar[621] := WCHAR#' ';
   SendWChar[622] := WCHAR#' ';
   SendWChar[623] := WCHAR#' ';
   SendWChar[624] := WCHAR#' ';
   SendWChar[625] := WCHAR#' ';
   SendWChar[626] := WCHAR#' ';
   SendWChar[627] := WCHAR#' ';
   SendWChar[628] := WCHAR#' ';
   SendWChar[629] := WCHAR#' ';
   SendWChar[630] := WCHAR#' ';
   SendWChar[631] := WCHAR#' ';
   SendWChar[632] := WCHAR#' ';
   SendWChar[633] := WCHAR#' ';
   SendWChar[634] := WCHAR#' ';
   SendWChar[635] := WCHAR#' ';
   SendWChar[636] := WCHAR#' ';
   SendWChar[637] := WCHAR#' ';
   SendWChar[638] := WCHAR#' ';
   SendWChar[639] := WCHAR#' ';
   SendWChar[640] := WCHAR#' ';
   SendWChar[641] := WCHAR#' ';
   SendWChar[642] := WCHAR#' ';
   SendWChar[643] := WCHAR#' ';
   SendWChar[644] := WCHAR#' ';
   SendWChar[645] := WCHAR#' ';
   SendWChar[646] := WCHAR#' ';
   SendWChar[647] := WCHAR#' ';
   SendWChar[648] := WCHAR#' ';
   SendWChar[649] := WCHAR#' ';
   SendWChar[650] := WCHAR#' ';
   SendWChar[651] := WCHAR#' ';
   SendWChar[652] := WCHAR#' ';
   SendWChar[653] := WCHAR#' ';
   SendWChar[654] := WCHAR#' ';
   SendWChar[655] := WCHAR#' ';
   SendWChar[656] := WCHAR#' ';
   SendWChar[657] := WCHAR#' ';
   SendWChar[658] := WCHAR#' ';
   SendWChar[659] := WCHAR#' ';
   SendWChar[660] := WCHAR#' ';
   SendWChar[661] := WCHAR#' ';
   SendWChar[662] := WCHAR#' ';
   SendWChar[663] := WCHAR#' ';
   SendWChar[664] := WCHAR#' ';
   SendWChar[665] := WCHAR#' ';
   SendWChar[666] := WCHAR#' ';
   SendWChar[667] := WCHAR#' ';
   SendWChar[668] := WCHAR#' ';
   SendWChar[669] := WCHAR#' ';
   SendWChar[670] := WCHAR#' ';
   SendWChar[671] := WCHAR#' ';
   SendWChar[672] := WCHAR#' ';
   SendWChar[673] := WCHAR#' ';
   SendWChar[674] := WCHAR#' ';
   SendWChar[675] := WCHAR#' ';
   SendWChar[676] := WCHAR#' ';
   SendWChar[677] := WCHAR#' ';
   SendWChar[678] := WCHAR#' ';
   SendWChar[679] := WCHAR#' ';
   SendWChar[680] := WCHAR#' ';
   SendWChar[681] := WCHAR#' ';
   SendWChar[682] := WCHAR#' ';
   SendWChar[683] := WCHAR#' ';
   SendWChar[684] := WCHAR#' ';
   SendWChar[685] := WCHAR#' ';
   SendWChar[686] := WCHAR#' ';
   SendWChar[687] := WCHAR#' ';
   SendWChar[688] := WCHAR#' ';
   SendWChar[689] := WCHAR#' ';
   SendWChar[690] := WCHAR#' ';
   SendWChar[691] := WCHAR#' ';
   SendWChar[692] := WCHAR#' ';
   SendWChar[693] := WCHAR#' ';
   SendWChar[694] := WCHAR#' ';
   SendWChar[695] := WCHAR#' ';
   SendWChar[696] := WCHAR#' ';
   SendWChar[697] := WCHAR#' ';
   SendWChar[698] := WCHAR#' ';
   SendWChar[699] := WCHAR#' ';
   SendWChar[700] := WCHAR#' ';
   SendWChar[701] := WCHAR#' ';
   SendWChar[702] := WCHAR#' ';
   SendWChar[703] := WCHAR#' ';
   SendWChar[704] := WCHAR#' ';
   SendWChar[705] := WCHAR#' ';
   SendWChar[706] := WCHAR#' ';
   SendWChar[707] := WCHAR#' ';
   SendWChar[708] := WCHAR#' ';
   SendWChar[709] := WCHAR#' ';
   SendWChar[710] := WCHAR#' ';
   SendWChar[711] := WCHAR#' ';
   SendWChar[712] := WCHAR#' ';
   SendWChar[713] := WCHAR#' ';
   SendWChar[714] := WCHAR#' ';
   SendWChar[715] := WCHAR#' ';
   SendWChar[716] := WCHAR#' ';
   SendWChar[717] := WCHAR#' ';
   SendWChar[718] := WCHAR#' ';
   SendWChar[719] := WCHAR#' ';
   SendWChar[720] := WCHAR#' ';
   SendWChar[721] := WCHAR#' ';
   SendWChar[722] := WCHAR#' ';
   SendWChar[723] := WCHAR#' ';
   SendWChar[724] := WCHAR#' ';
   SendWChar[725] := WCHAR#' ';
   SendWChar[726] := WCHAR#' ';
   SendWChar[727] := WCHAR#' ';
   SendWChar[728] := WCHAR#' ';
   SendWChar[729] := WCHAR#' ';
   SendWChar[730] := WCHAR#' ';
   SendWChar[731] := WCHAR#' ';
   SendWChar[732] := WCHAR#' ';
   SendWChar[733] := WCHAR#' ';
   SendWChar[734] := WCHAR#' ';
   SendWChar[735] := WCHAR#' ';
   SendWChar[736] := WCHAR#' ';
   SendWChar[737] := WCHAR#' ';
   SendWChar[738] := WCHAR#' ';
   SendWChar[739] := WCHAR#' ';
   SendWChar[740] := WCHAR#' ';
   SendWChar[741] := WCHAR#' ';
   SendWChar[742] := WCHAR#' ';
   SendWChar[743] := WCHAR#' ';
   SendWChar[744] := WCHAR#' ';
   SendWChar[745] := WCHAR#' ';
   SendWChar[746] := WCHAR#' ';
   SendWChar[747] := WCHAR#' ';
   SendWChar[748] := WCHAR#' ';
   SendWChar[749] := WCHAR#' ';
   SendWChar[750] := WCHAR#' ';
   SendWChar[751] := WCHAR#' ';
   SendWChar[752] := WCHAR#' ';
   SendWChar[753] := WCHAR#' ';
   SendWChar[754] := WCHAR#' ';
   SendWChar[755] := WCHAR#' ';
   SendWChar[756] := WCHAR#' ';
   SendWChar[757] := WCHAR#' ';
   SendWChar[758] := WCHAR#' ';
   SendWChar[759] := WCHAR#' ';
   SendWChar[760] := WCHAR#' ';
   SendWChar[761] := WCHAR#' ';
   SendWChar[762] := WCHAR#' ';
   SendWChar[763] := WCHAR#' ';
   SendWChar[764] := WCHAR#' ';
   SendWChar[765] := WCHAR#' ';
   SendWChar[766] := WCHAR#' ';
   SendWChar[767] := WCHAR#' ';
   SendWChar[768] := WCHAR#' ';
   SendWChar[769] := WCHAR#' ';
   SendWChar[770] := WCHAR#' ';
   SendWChar[771] := WCHAR#' ';
   SendWChar[772] := WCHAR#' ';
   SendWChar[773] := WCHAR#' ';
   SendWChar[774] := WCHAR#' ';
   SendWChar[775] := WCHAR#' ';
   SendWChar[776] := WCHAR#' ';
   SendWChar[777] := WCHAR#' ';
   SendWChar[778] := WCHAR#' ';
   SendWChar[779] := WCHAR#' ';
   SendWChar[780] := WCHAR#' ';
   SendWChar[781] := WCHAR#' ';
   SendWChar[782] := WCHAR#' ';
   SendWChar[783] := WCHAR#' ';
   SendWChar[784] := WCHAR#' ';
   SendWChar[785] := WCHAR#' ';
   SendWChar[786] := WCHAR#' ';
   SendWChar[787] := WCHAR#' ';
   SendWChar[788] := WCHAR#' ';
   SendWChar[789] := WCHAR#' ';
   SendWChar[790] := WCHAR#' ';
   SendWChar[791] := WCHAR#' ';
   SendWChar[792] := WCHAR#' ';
   SendWChar[793] := WCHAR#' ';
   SendWChar[794] := WCHAR#' ';
   SendWChar[795] := WCHAR#' ';
   SendWChar[796] := WCHAR#' ';
   SendWChar[797] := WCHAR#' ';
   SendWChar[798] := WCHAR#' ';
   SendWChar[799] := WCHAR#' ';
   SendWChar[800] := WCHAR#' ';
   SendWChar[801] := WCHAR#' ';
   SendWChar[802] := WCHAR#' ';
   SendWChar[803] := WCHAR#' ';
   SendWChar[804] := WCHAR#' ';
   SendWChar[805] := WCHAR#' ';
   SendWChar[806] := WCHAR#' ';
   SendWChar[807] := WCHAR#' ';
   SendWChar[808] := WCHAR#' ';
   SendWChar[809] := WCHAR#' ';